(* Logix 5000 project; controller PLC_MCC1201_220AP1 vendor 1 type 14 code 164 rev 35.11; software revision 35.00; part 17 of 25 *)
(* tags used below, declared in another part *)
   ACTIVE_MODE : ALIAS FOR N54[208].3;
   AFI : ALIAS FOR B3[7].15;
   B153 : DINT[20];
   B3 : DINT[102];
   BLOWER_ON : ALIAS FOR O[67].13;
   BRSH1_DN_FLT : ALIAS FOR I[43].1;
   BRSH1_DN_FWD : ALIAS FOR O[45].1;
   BRSH1_DN_SS2 : ALIAS FOR O[46].9;
   BRSH1_UP_FLT : ALIAS FOR I[43].0;
   BRSH1_UP_FWD : ALIAS FOR O[45].0;
   BRSH1_UP_SS2 : ALIAS FOR O[46].8;
   C2_NTH_IN_PE : ALIAS FOR N54[261].6;
   C2_NTH_IN_SS : ALIAS FOR N54[261].2;
   C2_NTH_OUT_PE : ALIAS FOR N54[261].5;
   C2_NTH_OUT_SS : ALIAS FOR N54[261].1;
   C2_STH_IN_PE : ALIAS FOR N54[261].8;
   C2_STH_IN_SS : ALIAS FOR N54[261].4;
   C2_STH_OUT_PE : ALIAS FOR N54[261].7;
   C2_STH_OUT_SS : ALIAS FOR N54[261].3;
   C3_ACTIVE_LAMP : ALIAS FOR N54[262].0;
   C5 : COUNTER[100];
   CBF_START_B : ALIAS FOR I[65].5;
   CBF_START_T : ALIAS FOR I[65].4;
   CBF_STOP_B : ALIAS FOR I[65].7;
   CBF_STOP_T : ALIAS FOR I[65].6;
   CHIP_BLOW_A : ALIAS FOR B3[1].3;
   CHIP_BLOW_M : ALIAS FOR B3[1].2;
   CR1_0FF_LAMP : ALIAS FOR O[67].9;
   CR1_AUTO : ALIAS FOR I[64].13;
   CR1_AUTO_MODE : ALIAS FOR N54[240].1;
   CR1_DOWN_PROX : ALIAS FOR I[64].11;
   CR1_DOWN_PWRLOS : ALIAS FOR N54[240].10;
   CR1_DOWN_RLY : ALIAS FOR O[67].1;
   CR1_DROP_COND : ALIAS FOR N54[240].13;
   CR1_DRV_FLT_LMP : ALIAS FOR O[66].8;
   CR1_DRV_FLT_RLY : ALIAS FOR O[66].9;
   CR1_DWN_PROX : ALIAS FOR N54[240].14;
   CR1_ESTOP : ALIAS FOR N54[240].3;
   CR1_FLT : ALIAS FOR I[65].0;
   CR1_FWD : ALIAS FOR O[66].0;
   CR1_MAN_MODE : ALIAS FOR N54[240].2;
   CR1_ON_LAMP : ALIAS FOR O[67].8;
   CR1_SS1 : ALIAS FOR O[66].2;
   CR1_START_PB : ALIAS FOR I[65].12;
   CR1_STOP_PB : ALIAS FOR I[65].13;
   CR1_TEST_PB : ALIAS FOR I[65].3;
   CR1_UP_PROX : ALIAS FOR I[64].12;
   CR1_UP_RLY : ALIAS FOR O[67].0;
   CR1_UPT_PROX : ALIAS FOR N54[240].15;
   ECLIPSE_OFF : ALIAS FOR N54[208].2;
   ECLIPSE_ON : ALIAS FOR N54[208].1;
   GENERATOR_ON : ALIAS FOR N54[240].11;
   GENERATOR_RUN : ALIAS FOR I[65].15;
   I : INT[128];
   M1_ALM_FLT_RLY : ALIAS FOR O[66].13;
   M1_DRV_CONT_ON : ALIAS FOR I[64].0;
   N128 : DINT[997];
   N163 : DINT[5];
   N164 : DINT[3];
   N53 : DINT[10];
   N54 : DINT[501];
   O : INT[128];
   RELDR_ESTOP : ALIAS FOR I[80].0;
   S : INT[128];
   SPNGE_DN_FLT : ALIAS FOR I[43].5;
   SPNGE_DN_FWD : ALIAS FOR O[45].5;
   SPNGE_DN_SS2 : ALIAS FOR O[46].13;
   SPNGE_UP_FLT : ALIAS FOR I[43].4;
   SPNGE_UP_FWD : ALIAS FOR O[45].4;
   SPNGE_UP_SS2 : ALIAS FOR O[46].12;
   Status : INT;   // INT tag to retrieve Status value through GSV created during conversion
   T4 : TIMER[100];
   T51 : TIMER[13];
   T57 : TIMER[100];
   VMCC_M1_RED : ALIAS FOR O[67].3;
   WASH_AK1_CR : ALIAS FOR N54[207].4;
   WASH_ARK_AUTO : ALIAS FOR N54[203].1;
   WASH_ARK_MANLMP : ALIAS FOR N54[203].9;
   WASH_ARK_MANUAL : ALIAS FOR N54[203].2;
   WASH_BR1_AUTO : ALIAS FOR N54[200].1;
   WASH_BR1_CR : ALIAS FOR N54[207].1;
   WASH_BR1_MANLMP : ALIAS FOR N54[200].9;
   WASH_BR1_MANUAL : ALIAS FOR N54[200].2;
   WASH_BR1_MOFF : ALIAS FOR N54[200].10;
   WASH_BR1_OFF : ALIAS FOR N54[200].4;
   WASH_BR1_ON : ALIAS FOR N54[200].3;
   WASH_BR1_SV : ALIAS FOR O[36].12;
   WASH_BR1LO_CON : ALIAS FOR N54[200].8;
   WASH_BR1LO_CVG : ALIAS FOR N54[206].1;
   WASH_BR1LO_RET : ALIAS FOR N54[200].7;
   WASH_BR1UP_CON : ALIAS FOR N54[200].6;
   WASH_BR1UP_CVG : ALIAS FOR N54[205].1;
   WASH_BR1UP_RET : ALIAS FOR N54[200].5;
   WASH_BR1UP_SV : ALIAS FOR O[36].14;
   WASH_BR2_CR : ALIAS FOR N54[207].2;
   WASH_CR_ACK : ALIAS FOR N54[207].0;
   WASH_CR_RESET : ALIAS FOR N54[207].7;
   WASH_SPG_AUTO : ALIAS FOR N54[202].1;
   WASH_SPG_CR : ALIAS FOR N54[207].3;
   WASH_SPG_MANLMP : ALIAS FOR N54[202].9;
   WASH_SPG_MANUAL : ALIAS FOR N54[202].2;
   WASH_SPG_MOFF : ALIAS FOR N54[202].10;
   WASH_SPG_OFF : ALIAS FOR N54[202].4;
   WASH_SPG_ON : ALIAS FOR N54[202].3;
   WASH_SPGLO_CON : ALIAS FOR N54[202].8;
   WASH_SPGLO_CVG : ALIAS FOR N54[206].3;
   WASH_SPGLO_RET : ALIAS FOR N54[202].7;
   WASH_SPGLO_SV : ALIAS FOR O[36].4;
   WASH_SPGUP_CON : ALIAS FOR N54[202].6;
   WASH_SPGUP_CVG : ALIAS FOR N54[205].3;
   WASH_SPGUP_RET : ALIAS FOR N54[202].5;
   WASH_SPGUP_SV : ALIAS FOR O[36].6;
(* MainProgram, continued *)

ROUTINE _46_NO1_CRUSH   (* ladder *)
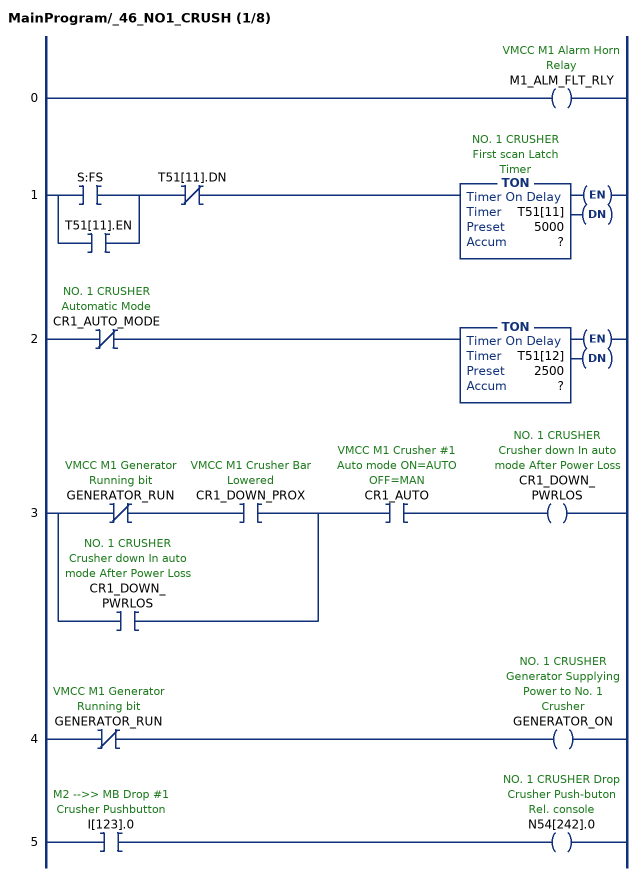
   0: OTE(M1_ALM_FLT_RLY);
   1: [XIC(S:FS) ,XIC(T51[11].EN) ]XIO(T51[11].DN)TON(T51[11],?,?);
   2: XIO(CR1_AUTO_MODE)TON(T51[12],?,?);
   3: [XIO(GENERATOR_RUN) XIC(CR1_DOWN_PROX) ,XIC(CR1_DOWN_PWRLOS) ]XIC(CR1_AUTO)OTE(CR1_DOWN_PWRLOS);
   4: XIO(GENERATOR_RUN)OTE(GENERATOR_ON);
   5: XIC(I[123].0)OTE(N54[242].0);
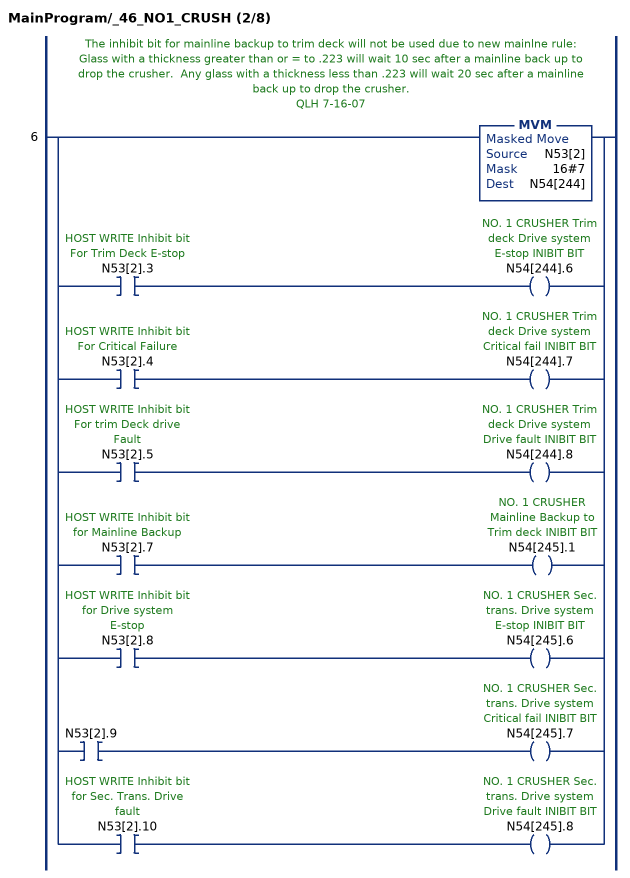
   // The inhibit bit for mainline backup to trim deck will not be used due to new mainlne rule:  Glass with a thickness greater than or = to .223 will wait 10 sec after a mainline back up to drop the crusher.  Any glass with a thickness less than .223 will wait 20 sec after a mainline back up to drop the crusher.
   // QLH 7-16-07
   6: [MVM(N53[2],16#7,N54[244]) ,XIC(N53[2].3) OTE(N54[244].6) ,XIC(N53[2].4) OTE(N54[244].7) ,XIC(N53[2].5) OTE(N54[244].8) ,XIC(N53[2].7) OTE(N54[245].1) ,XIC(N53[2].8) OTE(N54[245].6) ,XIC(N53[2].9) OTE(N54[245].7) ,XIC(N53[2].10) OTE(N54[245].8) ];
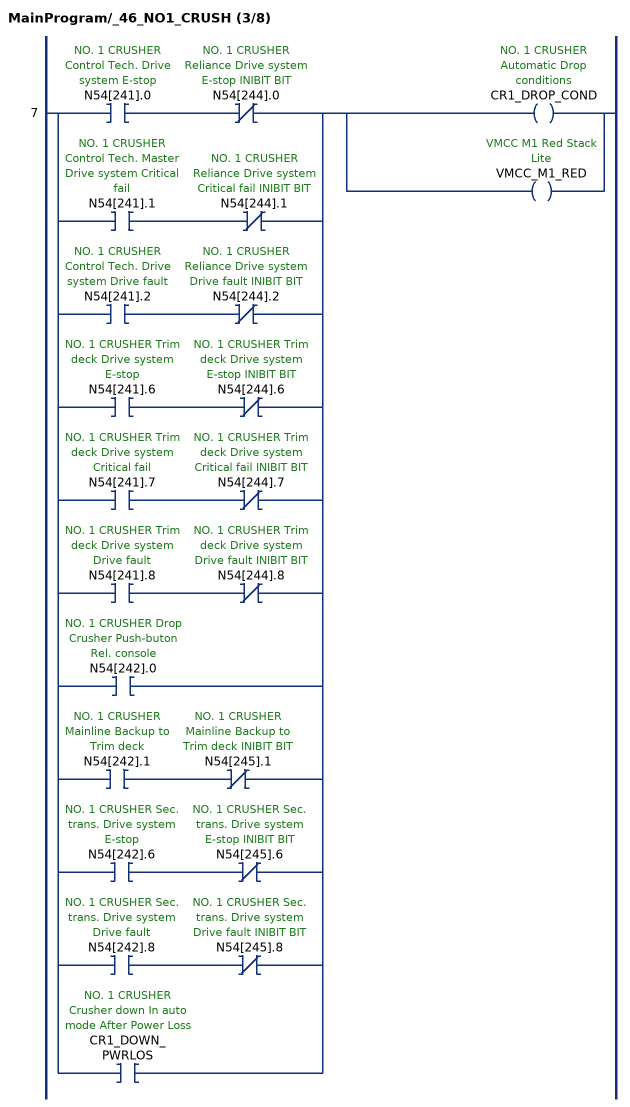
   7: [XIC(N54[241].0) XIO(N54[244].0) ,XIC(N54[241].1) XIO(N54[244].1) ,XIC(N54[241].2) XIO(N54[244].2) ,XIC(N54[241].6) XIO(N54[244].6) ,XIC(N54[241].7) XIO(N54[244].7) ,XIC(N54[241].8) XIO(N54[244].8) ,XIC(N54[242].0) ,XIC(N54[242].1) XIO(N54[245].1) ,XIC(N54[242].6) XIO(N54[245].6) ,XIC(N54[242].8) XIO(N54[245].8) ,XIC(CR1_DOWN_PWRLOS) ][OTE(CR1_DROP_COND) ,OTE(VMCC_M1_RED) ];
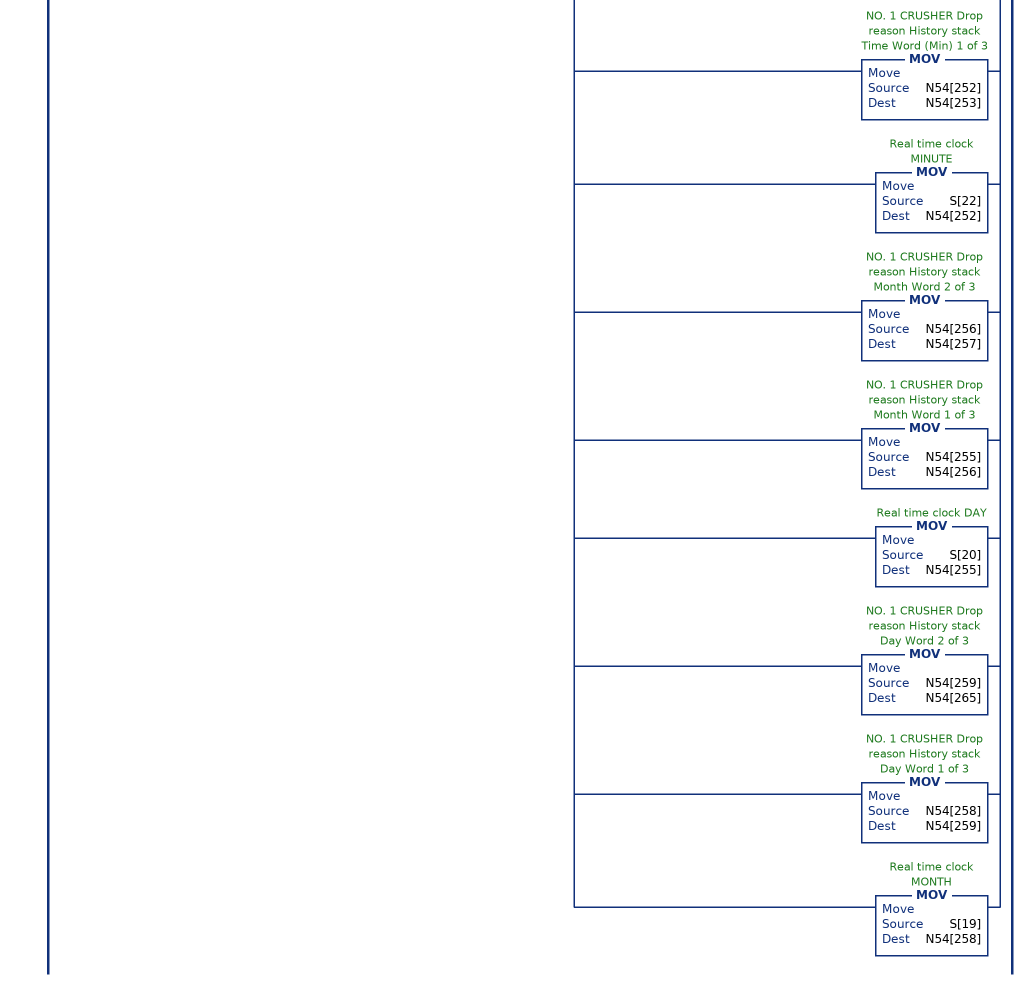
   // *** Generated by Migration Tool: Warning: Status files do not exist in RSLogix 5000. However this status file value is handled through the StatusFile routine. ***
   // *** Generated by Migration Tool: Warning: Status files do not exist in RSLogix 5000. However this status file value is handled through the StatusFile routine. ***
   // *** Generated by Migration Tool: Warning: Status files do not exist in RSLogix 5000. However this status file value is handled through the StatusFile routine. ***
   // *** Generated by Migration Tool: Warning: Status files do not exist in RSLogix 5000. However this status file value is handled through the StatusFile routine. ***
   8: XIC(CR1_DROP_COND)ONS(N54[240].8)XIO(CR1_DOWN_PROX)XIC(CR1_UP_PROX)[MOV(N54[247],N54[248]) ,MOV(N54[246],N54[247]) ,CLR(N54[246]) ,XIC(N54[241].0) XIO(N54[244].0) OTL(N54[246].0) ,XIC(N54[241].1) XIO(N54[244].1) OTL(N54[246].1) ,XIC(N54[241].2) XIO(N54[244].2) OTL(N54[246].2) ,XIC(N54[241].6) XIO(N54[244].6) OTL(N54[246].4) ,XIC(N54[241].7) XIO(N54[244].7) OTL(N54[246].5) ,XIC(N54[241].8) XIO(N54[244].8) OTL(N54[246].6) ,XIC(N54[242].0) OTL(N54[246].8) ,XIC(N54[242].1) XIO(N54[245].1) OTL(N54[246].9) ,XIC(N54[242].6) XIO(N54[245].6) OTL(N54[246].12) ,XIC(N54[242].8) XIO(N54[245].8) OTL(N54[246].14) ,XIC(CR1_DOWN_PWRLOS) OTL(N54[246].15) ,MOV(N54[250],N54[251]) ,MOV(N54[249],N54[250]) ,MOV(S[21],N54[249]) ,MOV(N54[253],N54[254]) ,MOV(N54[252],N54[253]) ,MOV(S[22],N54[252]) ,MOV(N54[256],N54[257]) ,MOV(N54[255],N54[256]) ,MOV(S[20],N54[255]) ,MOV(N54[259],N54[265]) ,MOV(N54[258],N54[259]) ,MOV(S[19],N54[258]) ];
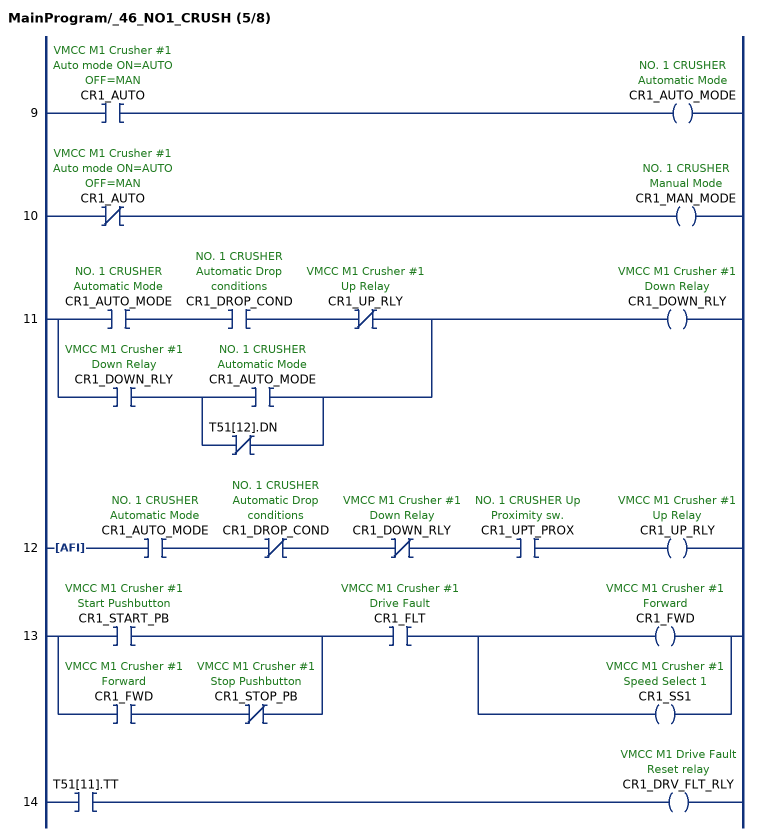
   9: XIC(CR1_AUTO)OTE(CR1_AUTO_MODE);
   10: XIO(CR1_AUTO)OTE(CR1_MAN_MODE);
   11: [XIC(CR1_AUTO_MODE) XIC(CR1_DROP_COND) XIO(CR1_UP_RLY) ,XIC(CR1_DOWN_RLY) [XIC(CR1_AUTO_MODE) ,XIO(T51[12].DN) ] ]OTE(CR1_DOWN_RLY);
   12: AFI()XIC(CR1_AUTO_MODE)XIO(CR1_DROP_COND)XIO(CR1_DOWN_RLY)XIC(CR1_UPT_PROX)OTE(CR1_UP_RLY);
   13: [XIC(CR1_START_PB) ,XIC(CR1_FWD) XIO(CR1_STOP_PB) ]XIC(CR1_FLT)[OTE(CR1_FWD) ,OTE(CR1_SS1) ];
   14: XIC(T51[11].TT)OTE(CR1_DRV_FLT_RLY);
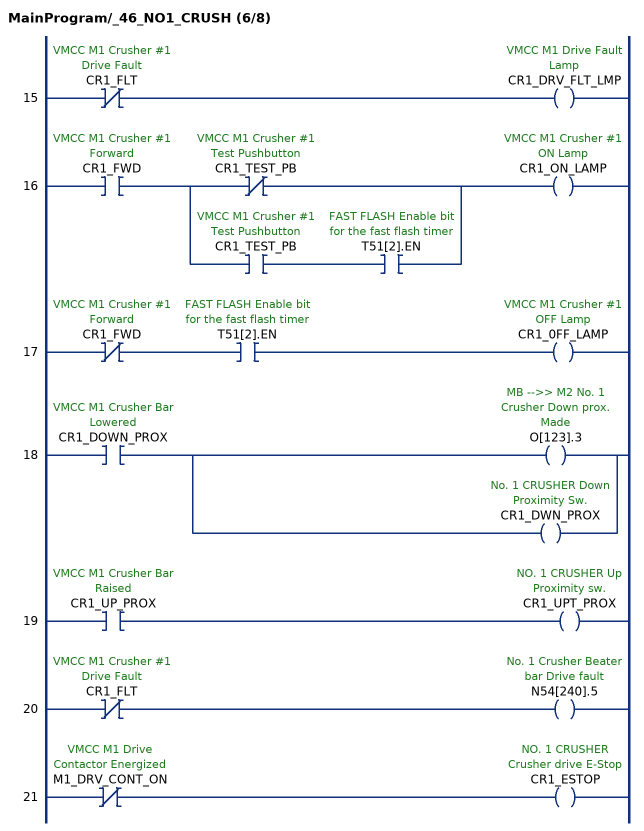
   15: XIO(CR1_FLT)OTE(CR1_DRV_FLT_LMP);
   16: XIC(CR1_FWD)[XIO(CR1_TEST_PB) ,XIC(CR1_TEST_PB) XIC(T51[2].EN) ]OTE(CR1_ON_LAMP);
   17: XIO(CR1_FWD)XIC(T51[2].EN)OTE(CR1_0FF_LAMP);
   18: XIC(CR1_DOWN_PROX)[OTE(O[123].3) ,OTE(CR1_DWN_PROX) ];
   19: XIC(CR1_UP_PROX)OTE(CR1_UPT_PROX);
   20: XIO(CR1_FLT)OTE(N54[240].5);
   21: XIO(M1_DRV_CONT_ON)OTE(CR1_ESTOP);
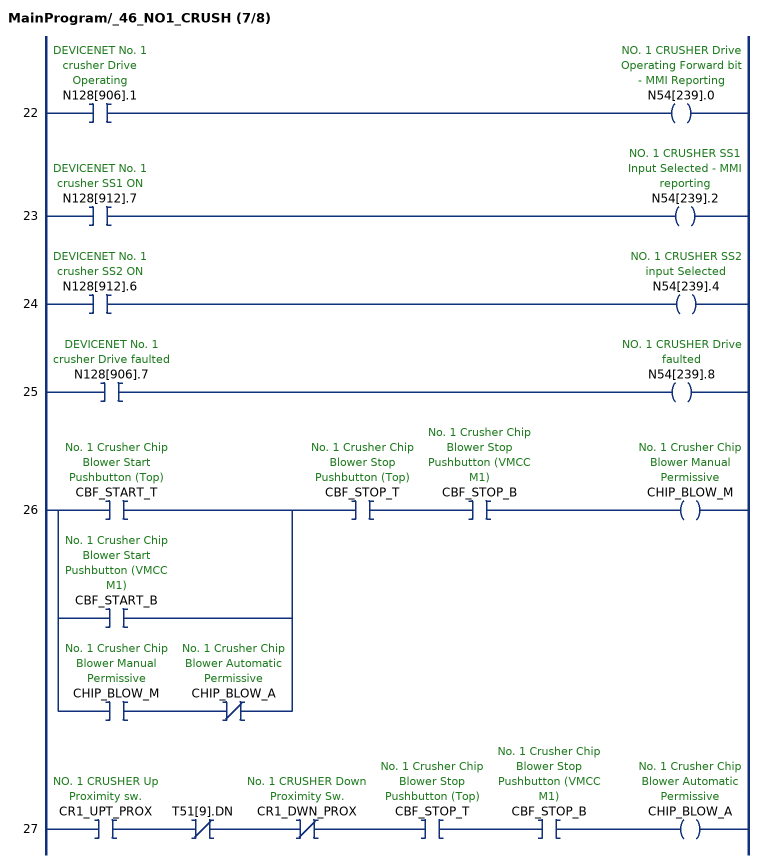
   22: XIC(N128[906].1)OTE(N54[239].0);
   23: XIC(N128[912].7)OTE(N54[239].2);
   24: XIC(N128[912].6)OTE(N54[239].4);
   25: XIC(N128[906].7)OTE(N54[239].8);
   26: [XIC(CBF_START_T) ,XIC(CBF_START_B) ,XIC(CHIP_BLOW_M) XIO(CHIP_BLOW_A) ]XIC(CBF_STOP_T)XIC(CBF_STOP_B)OTE(CHIP_BLOW_M);
   27: XIC(CR1_UPT_PROX)XIO(T51[9].DN)XIO(CR1_DWN_PROX)XIC(CBF_STOP_T)XIC(CBF_STOP_B)OTE(CHIP_BLOW_A);
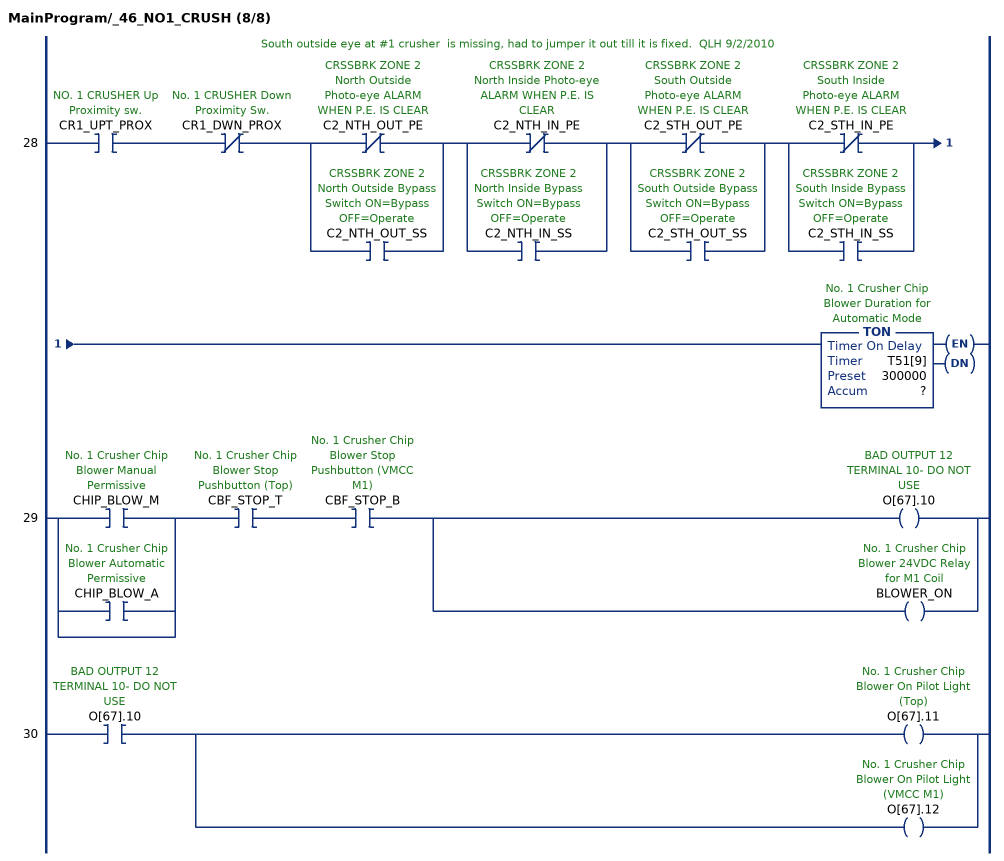
   // South outside eye at #1 crusher  is missing, had to jumper it out till it is fixed.  QLH 9/2/2010
   28: XIC(CR1_UPT_PROX)XIO(CR1_DWN_PROX)[XIO(C2_NTH_OUT_PE) ,XIC(C2_NTH_OUT_SS) ][XIO(C2_NTH_IN_PE) ,XIC(C2_NTH_IN_SS) ][XIO(C2_STH_OUT_PE) ,XIC(C2_STH_OUT_SS) ][XIO(C2_STH_IN_PE) ,XIC(C2_STH_IN_SS) ]TON(T51[9],?,?);
   29: [XIC(CHIP_BLOW_M) ,XIC(CHIP_BLOW_A) ,]XIC(CBF_STOP_T)XIC(CBF_STOP_B)[OTE(O[67].10) ,OTE(BLOWER_ON) ];
   30: XIC(O[67].10)[OTE(O[67].11) ,OTE(O[67].12) ];
END_ROUTINE

ROUTINE _47_WASHER   (* ladder *)
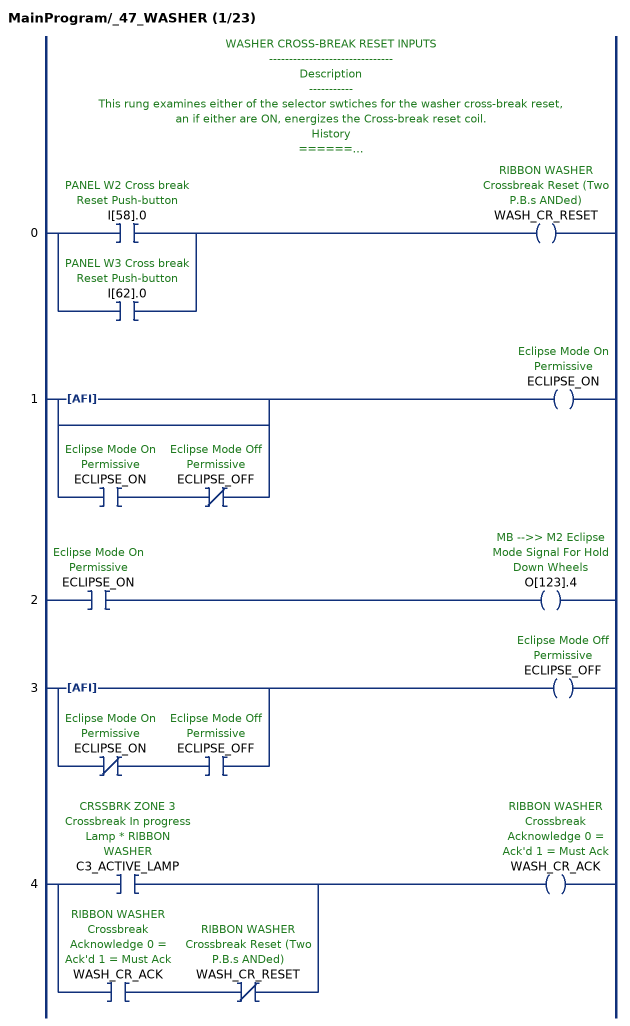
   // WASHER CROSS-BREAK RESET INPUTS
   // -------------------------------
   // Description
   // -----------
   // This rung examines either of the selector swtiches for the washer cross-break reset,
   // an if either are ON, energizes the Cross-break reset coil.
   // History
   // =======
   // DATE        DESCRIPTION                                              PROGRAMMER
   // ----        -----------                                              ----------
   // 1/29/96     Entered rung and coil comments.                          WAS
   0: [XIC(I[58].0) ,XIC(I[62].0) ]OTE(WASH_CR_RESET);
   1: [[AFI() ,] ,XIC(ECLIPSE_ON) XIO(ECLIPSE_OFF) ]OTE(ECLIPSE_ON);
   2: XIC(ECLIPSE_ON)OTE(O[123].4);
   3: [AFI() ,XIO(ECLIPSE_ON) XIC(ECLIPSE_OFF) ]OTE(ECLIPSE_OFF);
   4: [XIC(C3_ACTIVE_LAMP) ,XIC(WASH_CR_ACK) XIO(WASH_CR_RESET) ]OTE(WASH_CR_ACK);
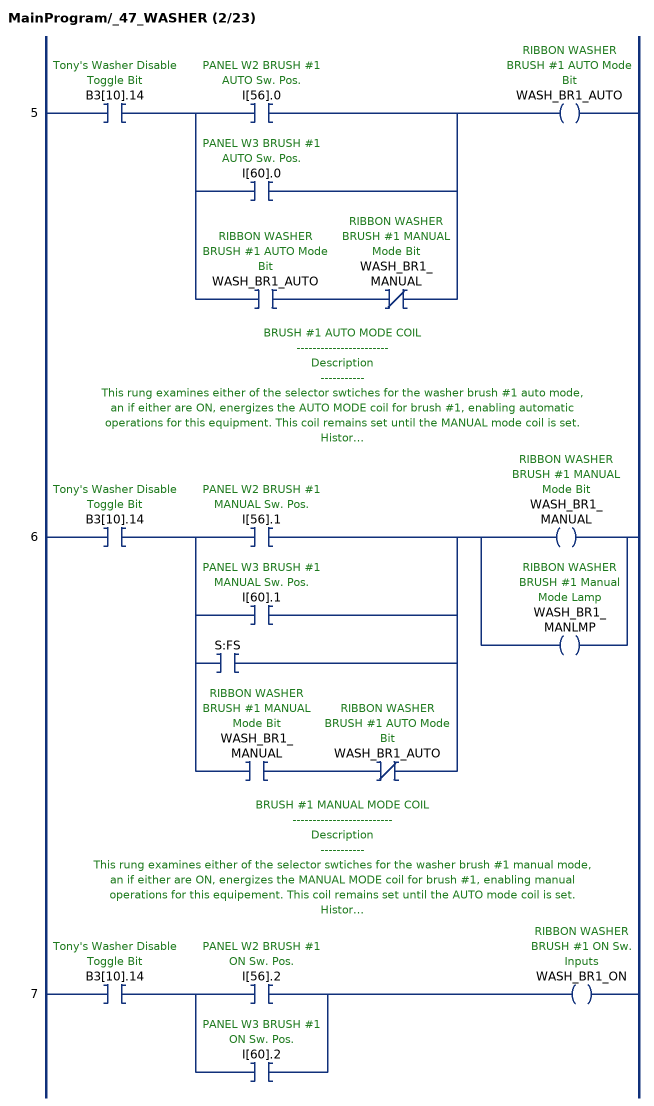
   5: XIC(B3[10].14)[[XIC(I[56].0) ,XIC(I[60].0) ] ,XIC(WASH_BR1_AUTO) XIO(WASH_BR1_MANUAL) ]OTE(WASH_BR1_AUTO);
   // BRUSH #1 AUTO MODE COIL
   // -----------------------
   // Description
   // -----------
   // This rung examines either of the selector swtiches for the washer brush #1 auto mode,
   // an if either are ON, energizes the AUTO MODE coil for brush #1, enabling automatic
   // operations for this equipment. This coil remains set until the MANUAL mode coil is set.
   // History
   // =======
   // DATE        DESCRIPTION                                              PROGRAMMER
   // ----        -----------                                              ----------
   // 1/29/96     Entered rung and coil comments.                          WAS
   6: XIC(B3[10].14)[[XIC(I[56].1) ,XIC(I[60].1) ,XIC(S:FS) ] ,XIC(WASH_BR1_MANUAL) XIO(WASH_BR1_AUTO) ][OTE(WASH_BR1_MANUAL) ,OTE(WASH_BR1_MANLMP) ];
   // BRUSH #1 MANUAL MODE COIL
   // -------------------------
   // Description
   // -----------
   // This rung examines either of the selector swtiches for the washer brush #1 manual mode,
   // an if either are ON, energizes the MANUAL MODE coil for brush #1, enabling manual
   // operations for this equipement. This coil remains set until the AUTO mode coil is set.
   // History
   // =======
   // DATE        DESCRIPTION                                              PROGRAMMER
   // ----        -----------                                              ----------
   // 1/29/96     Entered rung and coil comments.                          WAS
   7: XIC(B3[10].14)[XIC(I[56].2) ,XIC(I[60].2) ]OTE(WASH_BR1_ON);